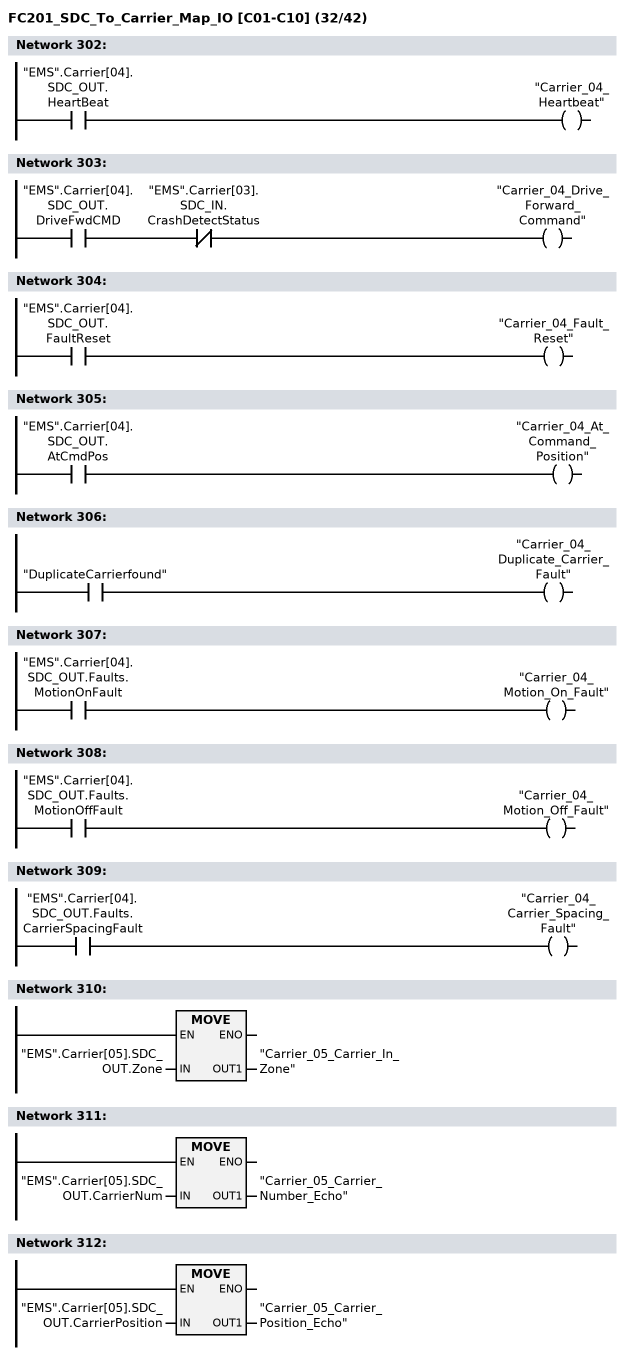
   RUNG wire#powerrail
      Contact( "EMS".Carrier[04].SDC_OUT.HeartBeat )
      Coil( "Carrier_04_Heartbeat" )
   END_RUNG
   // the same network as SCL:
   "Carrier_04_Heartbeat" := "EMS".Carrier[04].SDC_OUT.HeartBeat;
END_REGION

REGION Network 303
   RUNG wire#powerrail
      Contact( "EMS".Carrier[04].SDC_OUT.DriveFwdCMD )
      I_Contact( "EMS".Carrier[03].SDC_IN.CrashDetectStatus )
      Coil( "Carrier_04_Drive_Forward_Command" )
   END_RUNG
   // the same network as SCL:
   "Carrier_04_Drive_Forward_Command" := "EMS".Carrier[04].SDC_OUT.DriveFwdCMD AND NOT "EMS".Carrier[03].SDC_IN.CrashDetectStatus;
END_REGION

REGION Network 304
   RUNG wire#powerrail
      Contact( "EMS".Carrier[04].SDC_OUT.FaultReset )
      Coil( "Carrier_04_Fault_Reset" )
   END_RUNG
   // the same network as SCL:
   "Carrier_04_Fault_Reset" := "EMS".Carrier[04].SDC_OUT.FaultReset;
END_REGION

REGION Network 305
   RUNG wire#powerrail
      Contact( "EMS".Carrier[04].SDC_OUT.AtCmdPos )
      Coil( "Carrier_04_At_Command_Position" )
   END_RUNG
   // the same network as SCL:
   "Carrier_04_At_Command_Position" := "EMS".Carrier[04].SDC_OUT.AtCmdPos;
END_REGION

REGION Network 306
   RUNG wire#powerrail
      Contact( "DuplicateCarrierfound" )
      Coil( "Carrier_04_Duplicate_Carrier_Fault" )
   END_RUNG
   // the same network as SCL:
   "Carrier_04_Duplicate_Carrier_Fault" := "DuplicateCarrierfound";
END_REGION

REGION Network 307
   RUNG wire#powerrail
      Contact( "EMS".Carrier[04].SDC_OUT.Faults.MotionOnFault )
      Coil( "Carrier_04_Motion_On_Fault" )
   END_RUNG
   // the same network as SCL:
   "Carrier_04_Motion_On_Fault" := "EMS".Carrier[04].SDC_OUT.Faults.MotionOnFault;
END_REGION

REGION Network 308
   RUNG wire#powerrail
      Contact( "EMS".Carrier[04].SDC_OUT.Faults.MotionOffFault )
      Coil( "Carrier_04_Motion_Off_Fault" )
   END_RUNG
   // the same network as SCL:
   "Carrier_04_Motion_Off_Fault" := "EMS".Carrier[04].SDC_OUT.Faults.MotionOffFault;
END_REGION

REGION Network 309
   RUNG wire#powerrail
      Contact( "EMS".Carrier[04].SDC_OUT.Faults.CarrierSpacingFault )
      Coil( "Carrier_04_Carrier_Spacing_Fault" )
   END_RUNG
   // the same network as SCL:
   "Carrier_04_Carrier_Spacing_Fault" := "EMS".Carrier[04].SDC_OUT.Faults.CarrierSpacingFault;
END_REGION

REGION Network 310
   RUNG wire#powerrail
      Move(in := "EMS".Carrier[05].SDC_OUT.Zone, out1 => "Carrier_05_Carrier_In_Zone")
   END_RUNG
   // the same network as SCL:
   "Carrier_05_Carrier_In_Zone" := "EMS".Carrier[05].SDC_OUT.Zone;
END_REGION

REGION Network 311
   RUNG wire#powerrail
      Move(in := "EMS".Carrier[05].SDC_OUT.CarrierNum, out1 => "Carrier_05_Carrier_Number_Echo")
   END_RUNG
   // the same network as SCL:
   "Carrier_05_Carrier_Number_Echo" := "EMS".Carrier[05].SDC_OUT.CarrierNum;
END_REGION

REGION Network 312
   RUNG wire#powerrail
      Move(in := "EMS".Carrier[05].SDC_OUT.CarrierPosition, out1 => "Carrier_05_Carrier_Position_Echo")
   END_RUNG
   // the same network as SCL:
   "Carrier_05_Carrier_Position_Echo" := "EMS".Carrier[05].SDC_OUT.CarrierPosition;
END_REGION

REGION Network 313
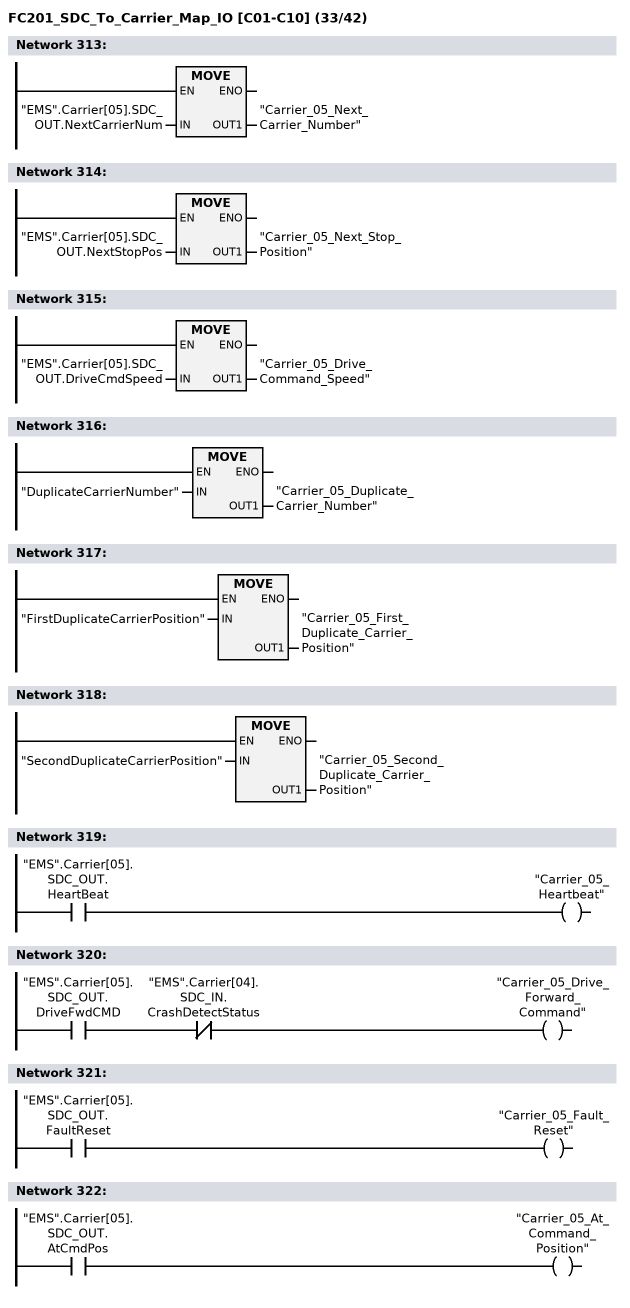
   RUNG wire#powerrail
      Move(in := "EMS".Carrier[05].SDC_OUT.NextCarrierNum, out1 => "Carrier_05_Next_Carrier_Number")
   END_RUNG
   // the same network as SCL:
   "Carrier_05_Next_Carrier_Number" := "EMS".Carrier[05].SDC_OUT.NextCarrierNum;
END_REGION

REGION Network 314
   RUNG wire#powerrail
      Move(in := "EMS".Carrier[05].SDC_OUT.NextStopPos, out1 => "Carrier_05_Next_Stop_Position")
   END_RUNG
   // the same network as SCL:
   "Carrier_05_Next_Stop_Position" := "EMS".Carrier[05].SDC_OUT.NextStopPos;
END_REGION

REGION Network 315
   RUNG wire#powerrail
      Move(in := "EMS".Carrier[05].SDC_OUT.DriveCmdSpeed, out1 => "Carrier_05_Drive_Command_Speed")
   END_RUNG
   // the same network as SCL:
   "Carrier_05_Drive_Command_Speed" := "EMS".Carrier[05].SDC_OUT.DriveCmdSpeed;
END_REGION

REGION Network 316
   RUNG wire#powerrail
      Move(in := "DuplicateCarrierNumber", out1 => "Carrier_05_Duplicate_Carrier_Number")
   END_RUNG
   // the same network as SCL:
   "Carrier_05_Duplicate_Carrier_Number" := "DuplicateCarrierNumber";
END_REGION

REGION Network 317
   RUNG wire#powerrail
      Move(in := "FirstDuplicateCarrierPosition", out1 => "Carrier_05_First_Duplicate_Carrier_Position")
   END_RUNG
   // the same network as SCL:
   "Carrier_05_First_Duplicate_Carrier_Position" := "FirstDuplicateCarrierPosition";
END_REGION

REGION Network 318
   RUNG wire#powerrail
      Move(in := "SecondDuplicateCarrierPosition", out1 => "Carrier_05_Second_Duplicate_Carrier_Position")
   END_RUNG
   // the same network as SCL:
   "Carrier_05_Second_Duplicate_Carrier_Position" := "SecondDuplicateCarrierPosition";
END_REGION

REGION Network 319
   RUNG wire#powerrail
      Contact( "EMS".Carrier[05].SDC_OUT.HeartBeat )
      Coil( "Carrier_05_Heartbeat" )
   END_RUNG
   // the same network as SCL:
   "Carrier_05_Heartbeat" := "EMS".Carrier[05].SDC_OUT.HeartBeat;
END_REGION

REGION Network 320
   RUNG wire#powerrail
      Contact( "EMS".Carrier[05].SDC_OUT.DriveFwdCMD )
      I_Contact( "EMS".Carrier[04].SDC_IN.CrashDetectStatus )
      Coil( "Carrier_05_Drive_Forward_Command" )
   END_RUNG
   // the same network as SCL:
   "Carrier_05_Drive_Forward_Command" := "EMS".Carrier[05].SDC_OUT.DriveFwdCMD AND NOT "EMS".Carrier[04].SDC_IN.CrashDetectStatus;
END_REGION

REGION Network 321
   RUNG wire#powerrail
      Contact( "EMS".Carrier[05].SDC_OUT.FaultReset )
      Coil( "Carrier_05_Fault_Reset" )
   END_RUNG
   // the same network as SCL:
   "Carrier_05_Fault_Reset" := "EMS".Carrier[05].SDC_OUT.FaultReset;
END_REGION

REGION Network 322
   RUNG wire#powerrail
      Contact( "EMS".Carrier[05].SDC_OUT.AtCmdPos )
      Coil( "Carrier_05_At_Command_Position" )
   END_RUNG
   // the same network as SCL:
   "Carrier_05_At_Command_Position" := "EMS".Carrier[05].SDC_OUT.AtCmdPos;
END_REGION

REGION Network 323
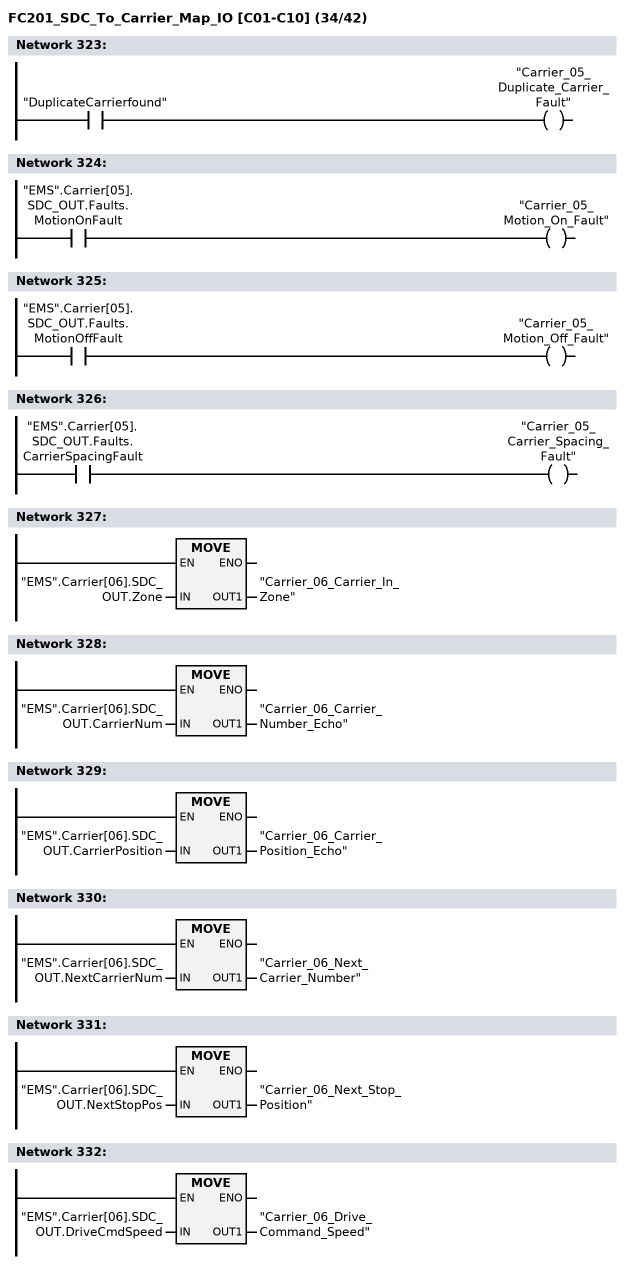
   RUNG wire#powerrail
      Contact( "DuplicateCarrierfound" )
      Coil( "Carrier_05_Duplicate_Carrier_Fault" )
   END_RUNG
   // the same network as SCL:
   "Carrier_05_Duplicate_Carrier_Fault" := "DuplicateCarrierfound";
END_REGION

REGION Network 324
   RUNG wire#powerrail
      Contact( "EMS".Carrier[05].SDC_OUT.Faults.MotionOnFault )
      Coil( "Carrier_05_Motion_On_Fault" )
   END_RUNG
   // the same network as SCL:
   "Carrier_05_Motion_On_Fault" := "EMS".Carrier[05].SDC_OUT.Faults.MotionOnFault;
END_REGION

REGION Network 325
   RUNG wire#powerrail
      Contact( "EMS".Carrier[05].SDC_OUT.Faults.MotionOffFault )
      Coil( "Carrier_05_Motion_Off_Fault" )
   END_RUNG
   // the same network as SCL:
   "Carrier_05_Motion_Off_Fault" := "EMS".Carrier[05].SDC_OUT.Faults.MotionOffFault;
END_REGION

REGION Network 326
   RUNG wire#powerrail
      Contact( "EMS".Carrier[05].SDC_OUT.Faults.CarrierSpacingFault )
      Coil( "Carrier_05_Carrier_Spacing_Fault" )
   END_RUNG
   // the same network as SCL:
   "Carrier_05_Carrier_Spacing_Fault" := "EMS".Carrier[05].SDC_OUT.Faults.CarrierSpacingFault;
END_REGION

REGION Network 327
   RUNG wire#powerrail
      Move(in := "EMS".Carrier[06].SDC_OUT.Zone, out1 => "Carrier_06_Carrier_In_Zone")
   END_RUNG
   // the same network as SCL:
   "Carrier_06_Carrier_In_Zone" := "EMS".Carrier[06].SDC_OUT.Zone;
END_REGION

REGION Network 328
   RUNG wire#powerrail
      Move(in := "EMS".Carrier[06].SDC_OUT.CarrierNum, out1 => "Carrier_06_Carrier_Number_Echo")
   END_RUNG
   // the same network as SCL:
   "Carrier_06_Carrier_Number_Echo" := "EMS".Carrier[06].SDC_OUT.CarrierNum;
END_REGION

REGION Network 329
   RUNG wire#powerrail
      Move(in := "EMS".Carrier[06].SDC_OUT.CarrierPosition, out1 => "Carrier_06_Carrier_Position_Echo")
   END_RUNG
   // the same network as SCL:
   "Carrier_06_Carrier_Position_Echo" := "EMS".Carrier[06].SDC_OUT.CarrierPosition;
END_REGION

REGION Network 330
   RUNG wire#powerrail
      Move(in := "EMS".Carrier[06].SDC_OUT.NextCarrierNum, out1 => "Carrier_06_Next_Carrier_Number")
   END_RUNG
   // the same network as SCL:
   "Carrier_06_Next_Carrier_Number" := "EMS".Carrier[06].SDC_OUT.NextCarrierNum;
END_REGION

REGION Network 331
   RUNG wire#powerrail
      Move(in := "EMS".Carrier[06].SDC_OUT.NextStopPos, out1 => "Carrier_06_Next_Stop_Position")
   END_RUNG
   // the same network as SCL:
   "Carrier_06_Next_Stop_Position" := "EMS".Carrier[06].SDC_OUT.NextStopPos;
END_REGION

REGION Network 332
   RUNG wire#powerrail
      Move(in := "EMS".Carrier[06].SDC_OUT.DriveCmdSpeed, out1 => "Carrier_06_Drive_Command_Speed")
   END_RUNG
   // the same network as SCL:
   "Carrier_06_Drive_Command_Speed" := "EMS".Carrier[06].SDC_OUT.DriveCmdSpeed;
END_REGION

REGION Network 333
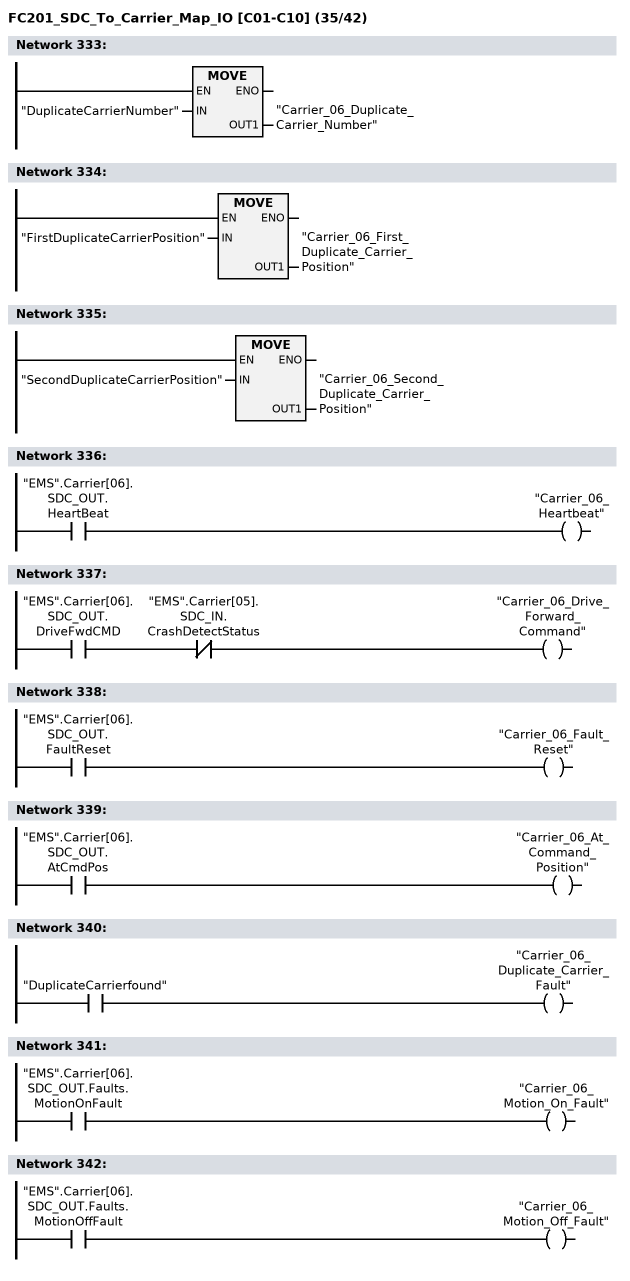
   RUNG wire#powerrail
      Move(in := "DuplicateCarrierNumber", out1 => "Carrier_06_Duplicate_Carrier_Number")
   END_RUNG
   // the same network as SCL:
   "Carrier_06_Duplicate_Carrier_Number" := "DuplicateCarrierNumber";
END_REGION

REGION Network 334
   RUNG wire#powerrail
      Move(in := "FirstDuplicateCarrierPosition", out1 => "Carrier_06_First_Duplicate_Carrier_Position")
   END_RUNG
   // the same network as SCL:
   "Carrier_06_First_Duplicate_Carrier_Position" := "FirstDuplicateCarrierPosition";
END_REGION

REGION Network 335
   RUNG wire#powerrail
      Move(in := "SecondDuplicateCarrierPosition", out1 => "Carrier_06_Second_Duplicate_Carrier_Position")
   END_RUNG
   // the same network as SCL:
   "Carrier_06_Second_Duplicate_Carrier_Position" := "SecondDuplicateCarrierPosition";
END_REGION

REGION Network 336
   RUNG wire#powerrail
      Contact( "EMS".Carrier[06].SDC_OUT.HeartBeat )
      Coil( "Carrier_06_Heartbeat" )
   END_RUNG
   // the same network as SCL:
   "Carrier_06_Heartbeat" := "EMS".Carrier[06].SDC_OUT.HeartBeat;
END_REGION

REGION Network 337
   RUNG wire#powerrail
      Contact( "EMS".Carrier[06].SDC_OUT.DriveFwdCMD )
      I_Contact( "EMS".Carrier[05].SDC_IN.CrashDetectStatus )
      Coil( "Carrier_06_Drive_Forward_Command" )
   END_RUNG
   // the same network as SCL:
   "Carrier_06_Drive_Forward_Command" := "EMS".Carrier[06].SDC_OUT.DriveFwdCMD AND NOT "EMS".Carrier[05].SDC_IN.CrashDetectStatus;
END_REGION

REGION Network 338
   RUNG wire#powerrail
      Contact( "EMS".Carrier[06].SDC_OUT.FaultReset )
      Coil( "Carrier_06_Fault_Reset" )
   END_RUNG
   // the same network as SCL:
   "Carrier_06_Fault_Reset" := "EMS".Carrier[06].SDC_OUT.FaultReset;
END_REGION

REGION Network 339
   RUNG wire#powerrail
      Contact( "EMS".Carrier[06].SDC_OUT.AtCmdPos )
      Coil( "Carrier_06_At_Command_Position" )
   END_RUNG
   // the same network as SCL:
   "Carrier_06_At_Command_Position" := "EMS".Carrier[06].SDC_OUT.AtCmdPos;
END_REGION

REGION Network 340
   RUNG wire#powerrail
      Contact( "DuplicateCarrierfound" )
      Coil( "Carrier_06_Duplicate_Carrier_Fault" )
   END_RUNG
   // the same network as SCL:
   "Carrier_06_Duplicate_Carrier_Fault" := "DuplicateCarrierfound";
END_REGION

REGION Network 341
   RUNG wire#powerrail
      Contact( "EMS".Carrier[06].SDC_OUT.Faults.MotionOnFault )
      Coil( "Carrier_06_Motion_On_Fault" )
   END_RUNG
   // the same network as SCL:
   "Carrier_06_Motion_On_Fault" := "EMS".Carrier[06].SDC_OUT.Faults.MotionOnFault;
END_REGION

REGION Network 342
   RUNG wire#powerrail
      Contact( "EMS".Carrier[06].SDC_OUT.Faults.MotionOffFault )
      Coil( "Carrier_06_Motion_Off_Fault" )
   END_RUNG
   // the same network as SCL:
   "Carrier_06_Motion_Off_Fault" := "EMS".Carrier[06].SDC_OUT.Faults.MotionOffFault;
END_REGION

REGION Network 343
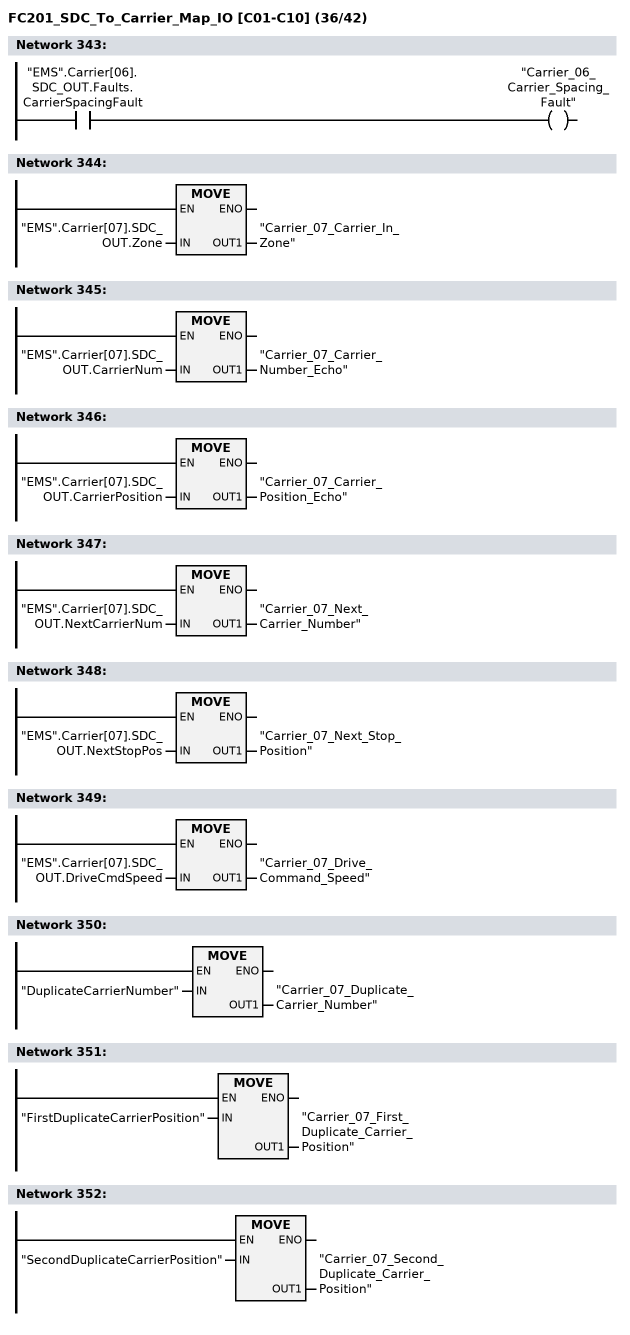
   RUNG wire#powerrail
      Contact( "EMS".Carrier[06].SDC_OUT.Faults.CarrierSpacingFault )
      Coil( "Carrier_06_Carrier_Spacing_Fault" )
   END_RUNG
   // the same network as SCL:
   "Carrier_06_Carrier_Spacing_Fault" := "EMS".Carrier[06].SDC_OUT.Faults.CarrierSpacingFault;
END_REGION

REGION Network 344
   RUNG wire#powerrail
      Move(in := "EMS".Carrier[07].SDC_OUT.Zone, out1 => "Carrier_07_Carrier_In_Zone")
   END_RUNG
   // the same network as SCL:
   "Carrier_07_Carrier_In_Zone" := "EMS".Carrier[07].SDC_OUT.Zone;
END_REGION

REGION Network 345
   RUNG wire#powerrail
      Move(in := "EMS".Carrier[07].SDC_OUT.CarrierNum, out1 => "Carrier_07_Carrier_Number_Echo")
   END_RUNG
   // the same network as SCL:
   "Carrier_07_Carrier_Number_Echo" := "EMS".Carrier[07].SDC_OUT.CarrierNum;
END_REGION

REGION Network 346
   RUNG wire#powerrail
      Move(in := "EMS".Carrier[07].SDC_OUT.CarrierPosition, out1 => "Carrier_07_Carrier_Position_Echo")
   END_RUNG
   // the same network as SCL:
   "Carrier_07_Carrier_Position_Echo" := "EMS".Carrier[07].SDC_OUT.CarrierPosition;
END_REGION

REGION Network 347
   RUNG wire#powerrail
      Move(in := "EMS".Carrier[07].SDC_OUT.NextCarrierNum, out1 => "Carrier_07_Next_Carrier_Number")
   END_RUNG
   // the same network as SCL:
   "Carrier_07_Next_Carrier_Number" := "EMS".Carrier[07].SDC_OUT.NextCarrierNum;
END_REGION

REGION Network 348
   RUNG wire#powerrail
      Move(in := "EMS".Carrier[07].SDC_OUT.NextStopPos, out1 => "Carrier_07_Next_Stop_Position")
   END_RUNG
   // the same network as SCL:
   "Carrier_07_Next_Stop_Position" := "EMS".Carrier[07].SDC_OUT.NextStopPos;
END_REGION

REGION Network 349
   RUNG wire#powerrail
      Move(in := "EMS".Carrier[07].SDC_OUT.DriveCmdSpeed, out1 => "Carrier_07_Drive_Command_Speed")
   END_RUNG
   // the same network as SCL:
   "Carrier_07_Drive_Command_Speed" := "EMS".Carrier[07].SDC_OUT.DriveCmdSpeed;
END_REGION

REGION Network 350
   RUNG wire#powerrail
      Move(in := "DuplicateCarrierNumber", out1 => "Carrier_07_Duplicate_Carrier_Number")
   END_RUNG
   // the same network as SCL:
   "Carrier_07_Duplicate_Carrier_Number" := "DuplicateCarrierNumber";
END_REGION

REGION Network 351
   RUNG wire#powerrail
      Move(in := "FirstDuplicateCarrierPosition", out1 => "Carrier_07_First_Duplicate_Carrier_Position")
   END_RUNG
   // the same network as SCL:
   "Carrier_07_First_Duplicate_Carrier_Position" := "FirstDuplicateCarrierPosition";
END_REGION

REGION Network 352
   RUNG wire#powerrail
      Move(in := "SecondDuplicateCarrierPosition", out1 => "Carrier_07_Second_Duplicate_Carrier_Position")
   END_RUNG
   // the same network as SCL:
   "Carrier_07_Second_Duplicate_Carrier_Position" := "SecondDuplicateCarrierPosition";
END_REGION

REGION Network 353
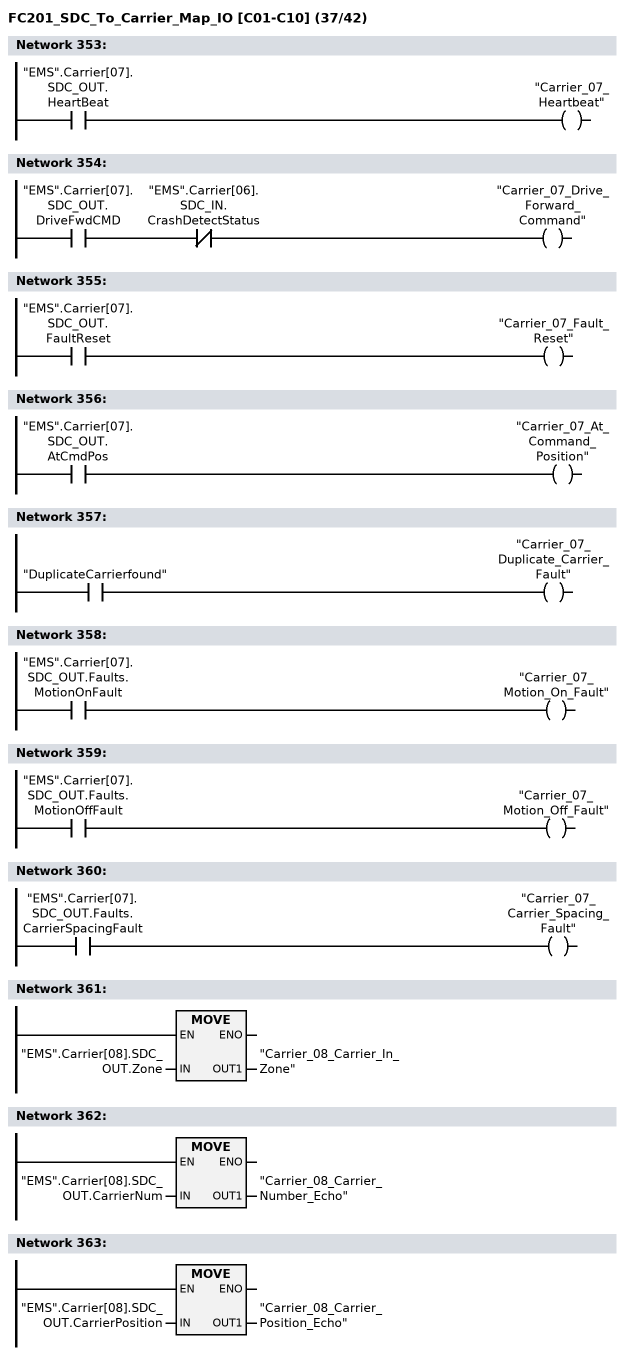
   RUNG wire#powerrail
      Contact( "EMS".Carrier[07].SDC_OUT.HeartBeat )
      Coil( "Carrier_07_Heartbeat" )
   END_RUNG
   // the same network as SCL:
   "Carrier_07_Heartbeat" := "EMS".Carrier[07].SDC_OUT.HeartBeat;
END_REGION

REGION Network 354
   RUNG wire#powerrail
      Contact( "EMS".Carrier[07].SDC_OUT.DriveFwdCMD )
      I_Contact( "EMS".Carrier[06].SDC_IN.CrashDetectStatus )
      Coil( "Carrier_07_Drive_Forward_Command" )
   END_RUNG
   // the same network as SCL:
   "Carrier_07_Drive_Forward_Command" := "EMS".Carrier[07].SDC_OUT.DriveFwdCMD AND NOT "EMS".Carrier[06].SDC_IN.CrashDetectStatus;
END_REGION

REGION Network 355
   RUNG wire#powerrail
      Contact( "EMS".Carrier[07].SDC_OUT.FaultReset )
      Coil( "Carrier_07_Fault_Reset" )
   END_RUNG
   // the same network as SCL:
   "Carrier_07_Fault_Reset" := "EMS".Carrier[07].SDC_OUT.FaultReset;
END_REGION

REGION Network 356
   RUNG wire#powerrail
      Contact( "EMS".Carrier[07].SDC_OUT.AtCmdPos )
      Coil( "Carrier_07_At_Command_Position" )
   END_RUNG
   // the same network as SCL:
   "Carrier_07_At_Command_Position" := "EMS".Carrier[07].SDC_OUT.AtCmdPos;
END_REGION

REGION Network 357
   RUNG wire#powerrail
      Contact( "DuplicateCarrierfound" )
      Coil( "Carrier_07_Duplicate_Carrier_Fault" )
   END_RUNG
   // the same network as SCL:
   "Carrier_07_Duplicate_Carrier_Fault" := "DuplicateCarrierfound";
END_REGION

REGION Network 358
   RUNG wire#powerrail
      Contact( "EMS".Carrier[07].SDC_OUT.Faults.MotionOnFault )
      Coil( "Carrier_07_Motion_On_Fault" )
   END_RUNG
   // the same network as SCL:
   "Carrier_07_Motion_On_Fault" := "EMS".Carrier[07].SDC_OUT.Faults.MotionOnFault;
END_REGION

REGION Network 359
   RUNG wire#powerrail
      Contact( "EMS".Carrier[07].SDC_OUT.Faults.MotionOffFault )
      Coil( "Carrier_07_Motion_Off_Fault" )
   END_RUNG
   // the same network as SCL:
   "Carrier_07_Motion_Off_Fault" := "EMS".Carrier[07].SDC_OUT.Faults.MotionOffFault;
END_REGION

REGION Network 360
   RUNG wire#powerrail
      Contact( "EMS".Carrier[07].SDC_OUT.Faults.CarrierSpacingFault )
      Coil( "Carrier_07_Carrier_Spacing_Fault" )
   END_RUNG
   // the same network as SCL:
   "Carrier_07_Carrier_Spacing_Fault" := "EMS".Carrier[07].SDC_OUT.Faults.CarrierSpacingFault;
END_REGION

REGION Network 361
   RUNG wire#powerrail
      Move(in := "EMS".Carrier[08].SDC_OUT.Zone, out1 => "Carrier_08_Carrier_In_Zone")
   END_RUNG
   // the same network as SCL:
   "Carrier_08_Carrier_In_Zone" := "EMS".Carrier[08].SDC_OUT.Zone;
END_REGION

REGION Network 362
   RUNG wire#powerrail
      Move(in := "EMS".Carrier[08].SDC_OUT.CarrierNum, out1 => "Carrier_08_Carrier_Number_Echo")
   END_RUNG
   // the same network as SCL:
   "Carrier_08_Carrier_Number_Echo" := "EMS".Carrier[08].SDC_OUT.CarrierNum;
END_REGION

REGION Network 363
   RUNG wire#powerrail
      Move(in := "EMS".Carrier[08].SDC_OUT.CarrierPosition, out1 => "Carrier_08_Carrier_Position_Echo")
   END_RUNG
   // the same network as SCL:
   "Carrier_08_Carrier_Position_Echo" := "EMS".Carrier[08].SDC_OUT.CarrierPosition;
END_REGION

REGION Network 364
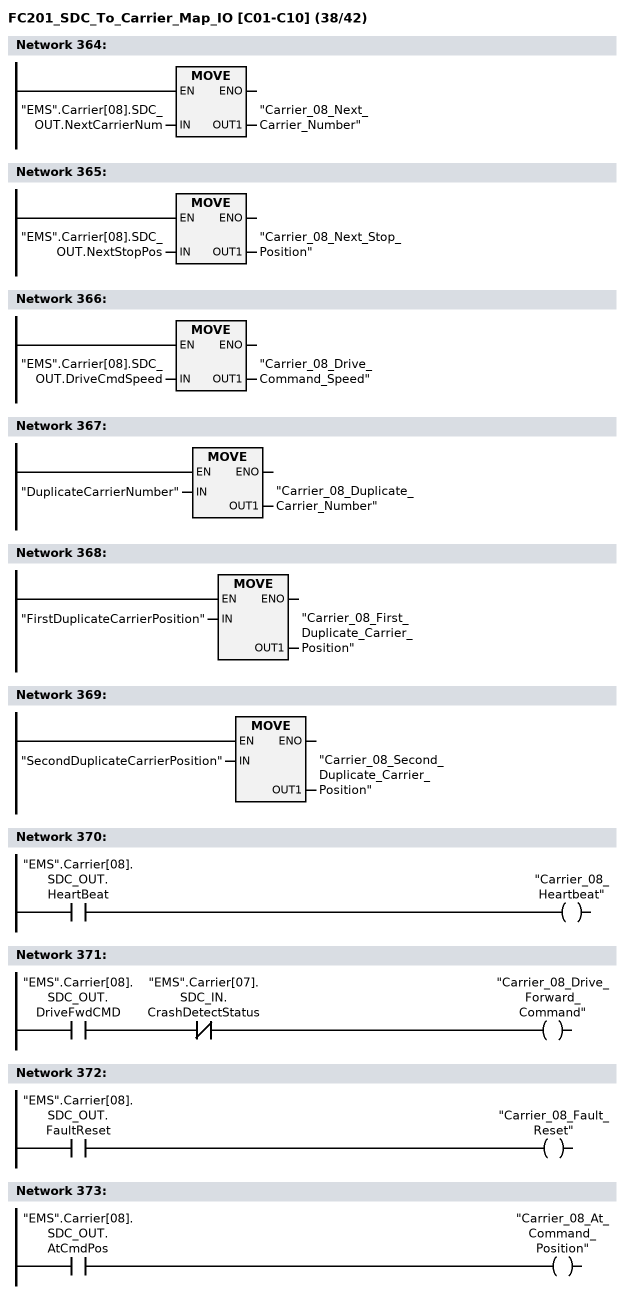
   RUNG wire#powerrail
      Move(in := "EMS".Carrier[08].SDC_OUT.NextCarrierNum, out1 => "Carrier_08_Next_Carrier_Number")
   END_RUNG
   // the same network as SCL:
   "Carrier_08_Next_Carrier_Number" := "EMS".Carrier[08].SDC_OUT.NextCarrierNum;
END_REGION

REGION Network 365
   RUNG wire#powerrail
      Move(in := "EMS".Carrier[08].SDC_OUT.NextStopPos, out1 => "Carrier_08_Next_Stop_Position")
   END_RUNG
   // the same network as SCL:
   "Carrier_08_Next_Stop_Position" := "EMS".Carrier[08].SDC_OUT.NextStopPos;
END_REGION

REGION Network 366
   RUNG wire#powerrail
      Move(in := "EMS".Carrier[08].SDC_OUT.DriveCmdSpeed, out1 => "Carrier_08_Drive_Command_Speed")
   END_RUNG
   // the same network as SCL:
   "Carrier_08_Drive_Command_Speed" := "EMS".Carrier[08].SDC_OUT.DriveCmdSpeed;
END_REGION

REGION Network 367
   RUNG wire#powerrail
      Move(in := "DuplicateCarrierNumber", out1 => "Carrier_08_Duplicate_Carrier_Number")
   END_RUNG
   // the same network as SCL:
   "Carrier_08_Duplicate_Carrier_Number" := "DuplicateCarrierNumber";
END_REGION

REGION Network 368
   RUNG wire#powerrail
      Move(in := "FirstDuplicateCarrierPosition", out1 => "Carrier_08_First_Duplicate_Carrier_Position")
   END_RUNG
   // the same network as SCL:
   "Carrier_08_First_Duplicate_Carrier_Position" := "FirstDuplicateCarrierPosition";
END_REGION

REGION Network 369
   RUNG wire#powerrail
      Move(in := "SecondDuplicateCarrierPosition", out1 => "Carrier_08_Second_Duplicate_Carrier_Position")
   END_RUNG
   // the same network as SCL:
   "Carrier_08_Second_Duplicate_Carrier_Position" := "SecondDuplicateCarrierPosition";
END_REGION

REGION Network 370
   RUNG wire#powerrail
      Contact( "EMS".Carrier[08].SDC_OUT.HeartBeat )
      Coil( "Carrier_08_Heartbeat" )
   END_RUNG
   // the same network as SCL:
   "Carrier_08_Heartbeat" := "EMS".Carrier[08].SDC_OUT.HeartBeat;
END_REGION

REGION Network 371
   RUNG wire#powerrail
      Contact( "EMS".Carrier[08].SDC_OUT.DriveFwdCMD )
      I_Contact( "EMS".Carrier[07].SDC_IN.CrashDetectStatus )
      Coil( "Carrier_08_Drive_Forward_Command" )
   END_RUNG
   // the same network as SCL:
   "Carrier_08_Drive_Forward_Command" := "EMS".Carrier[08].SDC_OUT.DriveFwdCMD AND NOT "EMS".Carrier[07].SDC_IN.CrashDetectStatus;
END_REGION

REGION Network 372
   RUNG wire#powerrail
      Contact( "EMS".Carrier[08].SDC_OUT.FaultReset )
      Coil( "Carrier_08_Fault_Reset" )
   END_RUNG
   // the same network as SCL:
   "Carrier_08_Fault_Reset" := "EMS".Carrier[08].SDC_OUT.FaultReset;
END_REGION

REGION Network 373
   RUNG wire#powerrail
      Contact( "EMS".Carrier[08].SDC_OUT.AtCmdPos )
      Coil( "Carrier_08_At_Command_Position" )
   END_RUNG
   // the same network as SCL:
   "Carrier_08_At_Command_Position" := "EMS".Carrier[08].SDC_OUT.AtCmdPos;
END_REGION

REGION Network 374
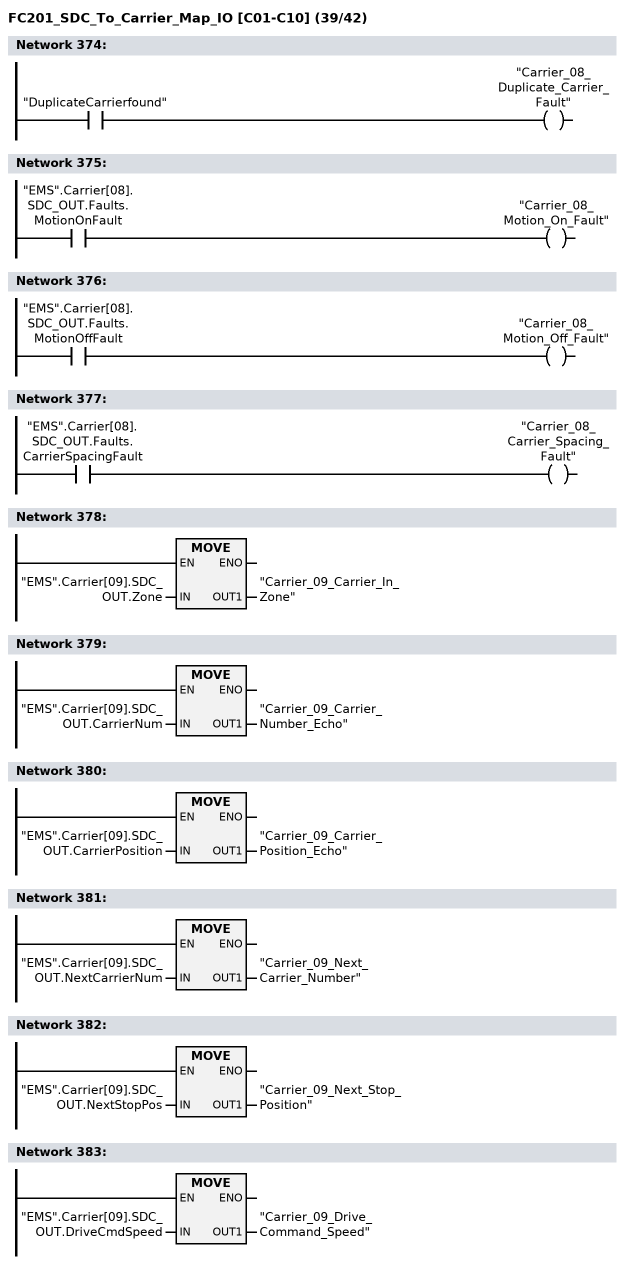
   RUNG wire#powerrail
      Contact( "DuplicateCarrierfound" )
      Coil( "Carrier_08_Duplicate_Carrier_Fault" )
   END_RUNG
   // the same network as SCL:
   "Carrier_08_Duplicate_Carrier_Fault" := "DuplicateCarrierfound";
END_REGION

REGION Network 375
   RUNG wire#powerrail
      Contact( "EMS".Carrier[08].SDC_OUT.Faults.MotionOnFault )
      Coil( "Carrier_08_Motion_On_Fault" )
   END_RUNG
   // the same network as SCL:
   "Carrier_08_Motion_On_Fault" := "EMS".Carrier[08].SDC_OUT.Faults.MotionOnFault;
END_REGION

REGION Network 376
   RUNG wire#powerrail
      Contact( "EMS".Carrier[08].SDC_OUT.Faults.MotionOffFault )
      Coil( "Carrier_08_Motion_Off_Fault" )
   END_RUNG
   // the same network as SCL:
   "Carrier_08_Motion_Off_Fault" := "EMS".Carrier[08].SDC_OUT.Faults.MotionOffFault;
END_REGION

REGION Network 377
   RUNG wire#powerrail
      Contact( "EMS".Carrier[08].SDC_OUT.Faults.CarrierSpacingFault )
      Coil( "Carrier_08_Carrier_Spacing_Fault" )
   END_RUNG
   // the same network as SCL:
   "Carrier_08_Carrier_Spacing_Fault" := "EMS".Carrier[08].SDC_OUT.Faults.CarrierSpacingFault;
END_REGION

REGION Network 378
   RUNG wire#powerrail
      Move(in := "EMS".Carrier[09].SDC_OUT.Zone, out1 => "Carrier_09_Carrier_In_Zone")
   END_RUNG
   // the same network as SCL:
   "Carrier_09_Carrier_In_Zone" := "EMS".Carrier[09].SDC_OUT.Zone;
END_REGION

REGION Network 379
   RUNG wire#powerrail
      Move(in := "EMS".Carrier[09].SDC_OUT.CarrierNum, out1 => "Carrier_09_Carrier_Number_Echo")
   END_RUNG
   // the same network as SCL:
   "Carrier_09_Carrier_Number_Echo" := "EMS".Carrier[09].SDC_OUT.CarrierNum;
END_REGION

REGION Network 380
   RUNG wire#powerrail
      Move(in := "EMS".Carrier[09].SDC_OUT.CarrierPosition, out1 => "Carrier_09_Carrier_Position_Echo")
   END_RUNG
   // the same network as SCL:
   "Carrier_09_Carrier_Position_Echo" := "EMS".Carrier[09].SDC_OUT.CarrierPosition;
END_REGION

REGION Network 381
   RUNG wire#powerrail
      Move(in := "EMS".Carrier[09].SDC_OUT.NextCarrierNum, out1 => "Carrier_09_Next_Carrier_Number")
   END_RUNG
   // the same network as SCL:
   "Carrier_09_Next_Carrier_Number" := "EMS".Carrier[09].SDC_OUT.NextCarrierNum;
END_REGION

REGION Network 382
   RUNG wire#powerrail
      Move(in := "EMS".Carrier[09].SDC_OUT.NextStopPos, out1 => "Carrier_09_Next_Stop_Position")
   END_RUNG
   // the same network as SCL:
   "Carrier_09_Next_Stop_Position" := "EMS".Carrier[09].SDC_OUT.NextStopPos;
END_REGION

REGION Network 383
   RUNG wire#powerrail
      Move(in := "EMS".Carrier[09].SDC_OUT.DriveCmdSpeed, out1 => "Carrier_09_Drive_Command_Speed")
   END_RUNG
   // the same network as SCL:
   "Carrier_09_Drive_Command_Speed" := "EMS".Carrier[09].SDC_OUT.DriveCmdSpeed;
END_REGION

REGION Network 384
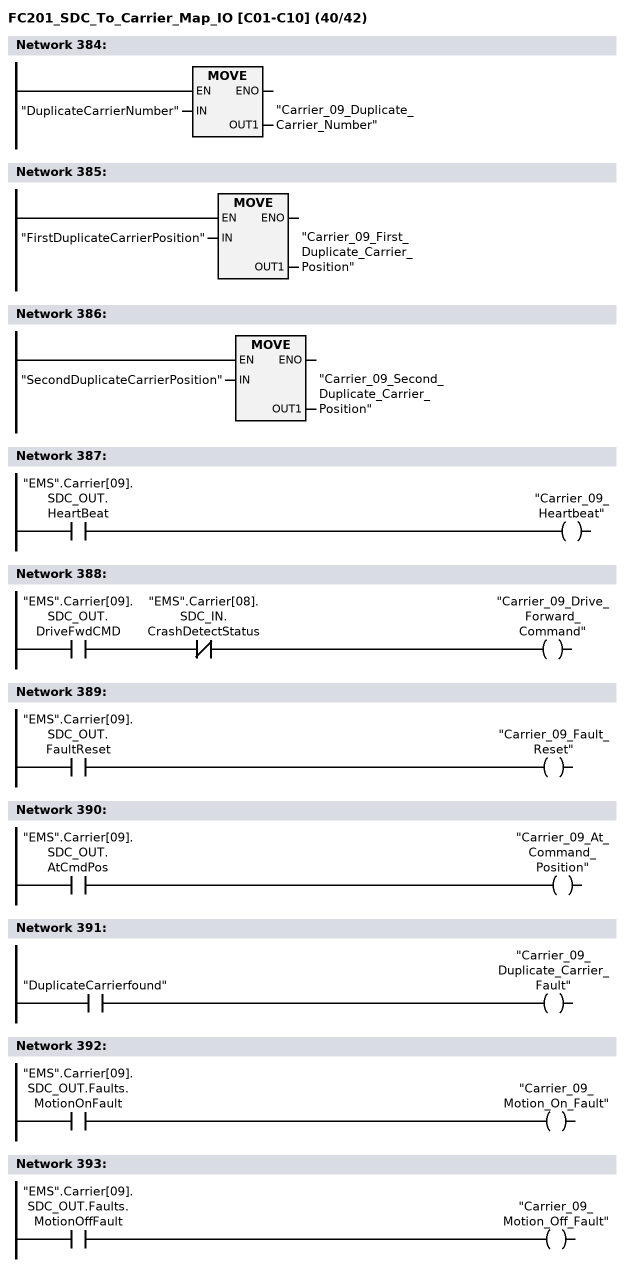
   RUNG wire#powerrail
      Move(in := "DuplicateCarrierNumber", out1 => "Carrier_09_Duplicate_Carrier_Number")
   END_RUNG
   // the same network as SCL:
   "Carrier_09_Duplicate_Carrier_Number" := "DuplicateCarrierNumber";
END_REGION
